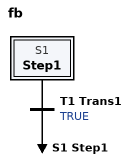
   // sequencer 1
   INITIAL_STEP Step1:   // S1, max time T#10S, warning time T#7S
   END_STEP
   TRANSITION Trans1 FROM Step1 TO Step1   // T1, jump
      := TRUE;
   END_TRANSITION
END_FUNCTION_BLOCK

ORGANIZATION_BLOCK "Main"   // OB1, LAD, ProgramCycle
TITLE = "Main Program Sweep (Cycle)"
{ S7_Optimized_Access := 'TRUE' }
VERSION : 0.1
   VAR_INPUT
      Initial_Call : Bool;   // Initial call of this OB
      Remanence : Bool;   // =True, if remanent data are available
   END_VAR
BEGIN

REGION Network 1
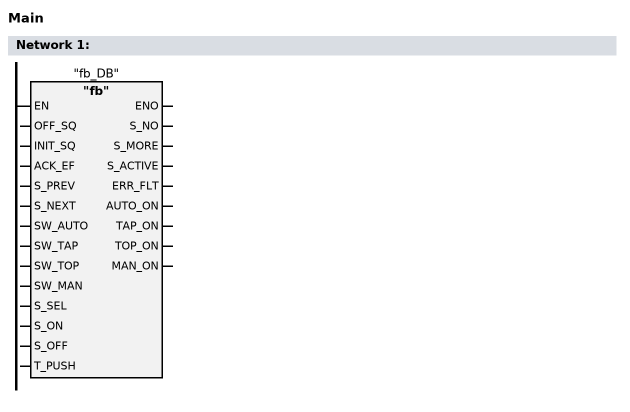
   RUNG wire#powerrail
      "fb_DB"(OFF_SQ :=, INIT_SQ :=, ACK_EF :=, S_PREV :=, S_NEXT :=, SW_AUTO :=, SW_TAP :=, SW_TOP :=, SW_MAN :=, S_SEL :=, S_ON :=, S_OFF :=, T_PUSH :=, S_NO =>, S_MORE =>, S_ACTIVE =>, ERR_FLT =>, AUTO_ON =>, TAP_ON =>, TOP_ON =>, MAN_ON =>)
   END_RUNG
   // the same network as SCL:
   "fb_DB"();   // "fb"
END_REGION
END_ORGANIZATION_BLOCK

(* ===== HMI "HMI_RT_2" =====
system functions are stored by id; their names below are inferred from use
connection "Connection_1": ETHERNET, SIMATIC S7 300/400 MPI
connection "HMI_Connection_1": ETHERNET, SIMATIC S7 300/400 MPI

HMI tags "Default tag table"
   "Tag_ScreenNumber" : UInt, internal
   "Greutate" : Int AT %DB7.DBW2, 1 s
   "LOAD" : Bool = PLC Banda_1_DB.Btn_LOAD AT %DB8.DBX0.4, 1 s
   "Manuala" : UInt, internal
   "Automata" : UInt, internal
   "StatieDistributie" : UInt, internal
   "StatieHidraulica" : UInt, internal
   "StatieIncarcare" : UInt, internal
   "Poz_Piston_1" : Int = PLC DB_general.Poz_Piston_1 AT %DB2.DBW2, 500 ms
   "Emg_Stop" : Bool = PLC Emg_Stop AT %I0.2, 1 s
   "Poz_Cutie" : Int = PLC Poz_Cutie AT %MW0, 500 ms
   "DB_general_Stare_Poz_Incarcare" : Bool = PLC DB_general.Stare_Poz_Incarcare AT %DB2.DBX0.0, 1 s
   "ON/OFF" : Bool = PLC "ON/OFF" AT %M2.1, 1 s
   "Viz_Cutie_Cursa_Scurta" : Bool = PLC Viz_Cutie_Cursa_Scurta AT %M2.2, 500 ms
   "Final_Cursa_P1" : Bool = PLC Final_Cursa_Piston_1 AT %M2.5, 1 s
   "Locuri_A" : Int = PLC DB_HMI.Locuri_A AT %DB19.DBW0, 1 s
   "Locuri_B" : Int = PLC DB_HMI.Locuri_B AT %DB19.DBW2, 1 s
   "Locuri_C" : Int = PLC DB_HMI.Locuri_C AT %DB19.DBW4, 1 s
   "Loc_Ocupat_A" : Int AT %DB1.DBW0, 1 s
   "DB_general_Poz_Piston_1" : Int = PLC DB_general.Poz_Piston_1 AT %DB2.DBW2, 1 s
   "DB_HMI_A_Pressed" : Bool = PLC DB_HMI.A_Pressed AT %DB19.DBX6.0, 1 s
   "DB_HMI_B_Pressed" : Bool = PLC DB_HMI.B_Pressed AT %DB19.DBX6.1, 1 s
   "DB_HMI_C_Pressed" : Bool = PLC DB_HMI.C_Pressed AT %DB19.DBX6.2, 1 s
   "DB_HMI_Cutie_Manuala" : Bool = PLC DB_HMI.Cutie_Manuala AT %DB19.DBX6.4, 1 s
   "DB_HMI_Cutie_Automata" : Bool = PLC DB_HMI.Cutie_Automata AT %DB19.DBX6.3, 1 s
   "DB_HMI_Viz_Cutie_Scurta" : Bool = PLC DB_HMI.Viz_Cutie_Scurta AT %DB19.DBX6.5, 1 s
   "DB_general_Senzor_1_Incarcare" : Bool = PLC DB_general.Senzor_1_Incarcare AT %DB2.DBX0.2, 1 s
   "DB_general_Senzor_2_Incarcare" : Bool = PLC DB_general.Senzor_2_Incarcare AT %DB2.DBX0.3, 1 s
   "DB_HMI_Tip_Cutie" : Int = PLC DB_HMI.Tip_Cutie_Lung AT %DB19.DBW8, 1 s
   "DB_HMI_LOAD" : Int = PLC DB_HMI.LOAD AT %DB19.DBW12, 1 s
   "DB_HMI_Transport" : Bool = PLC DB_HMI.Transport AT %DB19.DBX14.0, 1 s
   "DB_HMI_Viz_Cutie_Lunga" : Bool = PLC DB_HMI.Viz_Cutie_Lunga AT %DB19.DBX6.6, 1 s
   "DB_HMI_Tip_Cutie_Scurt" : Int = PLC DB_HMI.Tip_Cutie_Scurt AT %DB19.DBW10, 1 s
   "DB_general_Senzor_1_Descarcare" : Bool = PLC DB_general.Senzor_1_Descarcare AT %DB2.DBX0.4, 1 s
   "Stop" : Bool = PLC Stop AT %I0.1, 1 s
   "Start" : Bool = PLC Start AT %I0.0, 1 s
   "Man/Auto" : Bool = PLC "Man/Auto" AT %I0.3, 1 s
   "DB_general_Valoare" : Int = PLC DB_general.Valoare AT %DB2.DBW14, 1 s
   "DB_general_Piston_Cursa_Completa" : Int = PLC DB_general.Piston_1_Cursa_Completa AT %DB2.DBW16, 500 ms
   "DB_HMI_Viz_Cutie_Banda_1" : Bool = PLC DB_HMI.Viz_Cutie_Banda_1 AT %DB19.DBX14.2, 500 ms
   "DB_HMI_Ack_Load" : Bool = PLC DB_HMI.Ack_Load AT %DB19.DBX14.3, 1 s
   "DB_HMI_Piston_1_Status" : Int = PLC DB_HMI.Piston_1_Status AT %DB19.DBW16, 1 s
   "DB_HMI_Piston_2_Status" : Int = PLC DB_HMI.Piston_2_Status AT %DB19.DBW18, 1 s
   "DB_general_Piston_2_Cursa_Completa" : Int = PLC DB_general.Piston_2_Cursa_Completa AT %DB2.DBW18, 500 ms
   "DB_HMI_Load_RDY" : Bool = PLC DB_HMI.Load_RDY AT %DB19.DBX20.0, 1 s
   "DB_general_Poz_Cutie_Bile" : Int = PLC DB_general.Poz_Cutie_Bile AT %DB2.DBW8, 500 ms
   "DB_HMI_Viz_Cutie_A" : Bool = PLC DB_HMI.Viz_Cutie_A AT %DB19.DBX20.1, 1 s
   "DB_HMI_Viz_Cutie_B" : Bool = PLC DB_HMI.Viz_Cutie_B AT %DB19.DBX20.2, 1 s
   "DB_HMI_Viz_Cutie_C" : Bool = PLC DB_HMI.Viz_Cutie_C AT %DB19.DBX20.3, 1 s
   "DB_HMI_LOAD_A" : Bool = PLC DB_HMI.LOAD_A AT %DB19.DBX28.0, 1 s
   "DB_general_Piston_Incarcare_A" : Int = PLC DB_general.Piston_Incarcare_A AT %DB2.DBW30, 500 ms
   "DB_HMI_LOAD_B" : Bool = PLC DB_HMI.LOAD_B AT %DB19.DBX28.1, 1 s
   "DB_HMI_LOAD_C" : Bool = PLC DB_HMI.LOAD_C AT %DB19.DBX28.2, 1 s
   "DB_general_Piston_Incarcare_B" : Int = PLC DB_general.Piston_Incarcare_B AT %DB2.DBW32, 1 s
   "DB_general_Piston_Incarcare_C" : Int = PLC DB_general.Piston_Incarcare_C AT %DB2.DBW34, 1 s
   "DB_HMI_Status_Piston_A" : Int = PLC DB_HMI.Status_Piston_A AT %DB19.DBW22, 1 s
   "DB_HMI_Status_Piston_B" : Int = PLC DB_HMI.Status_Piston_B AT %DB19.DBW24, 1 s
   "DB_HMI_Status_Piston_C" : Int = PLC DB_HMI.Status_Piston_C AT %DB19.DBW26, 1 s
   "DB_HMI_Status_Banda_Bile" : Int = PLC DB_HMI.Status_Banda_Bile AT %DB19.DBW30, 1 s
   "DB_HMI_Sageata_Deplasare_Banda_Bile" : Bool = PLC DB_HMI.Sageata_Deplasare_Banda_Bile AT %DB19.DBX32.0, 1 s
   "DB_HMI_Temp_Ulei" : Int = PLC DB_HMI.Temp_Ulei AT %DB19.DBW34, 500 ms
   "DB_HMI_Volum_Ulei" : Int = PLC DB_HMI.Volum_Ulei AT %DB19.DBW40, 1 s
   "DB_HMI_Add_Ulei" : Bool = PLC DB_HMI.Add_Ulei AT %DB19.DBX42.0, 1 s
   "DB_HMI_Sub_Ulei" : Bool = PLC DB_HMI.Sub_Ulei AT %DB19.DBX42.1, 1 s
   "DB_HMI_Start_System" : Bool = PLC DB_HMI.Start_System AT %DB19.DBX42.2, 1 s
   "DB_HMI_Racire_Ulei" : Bool = PLC DB_HMI.Racire_Ulei AT %DB19.DBX42.3, 1 s
   "DB_HMI_Set_T0" : Bool = PLC DB_HMI.Set_T0 AT %DB19.DBX42.6, 1 s
   "DB_HMI_Set_T50" : Bool = PLC DB_HMI.Set_T50 AT %DB19.DBX42.7, 1 s
   "DB_HMI_START_SIM" : Bool = PLC DB_HMI.START_SIM AT %DB19.DBX43.0, 1 s
   "DB_SIM_BTN_RESET" : Bool = PLC DB_SIM.BTN_RESET AT %DB40.DBX0.4, 1 s
   "DB_HMI_TEST_LOAD" : Bool = PLC DB_HMI.BTN_LOAD AT %DB19.DBX43.1, 1 s
   "DB_Alarme_Emg_Stop" : Int = PLC DB_Alarme.Emg_Stop AT %DB46.DBW0, 1 s

discrete alarms
   1: 'Emergency Stop', class Errors, trigger "DB_Alarme_Emg_Stop" bit 0

analog alarms
   1: 'Limita greutate depasita / Gewichtslimit überschritten', class Warnings, trigger "Greutate"
   2: 'No more free spaces in A slot / Keine freien Plätze mehr im A-Steckplatz', class Acknowledgement, trigger "Locuri_A"
   3: 'No more free spaces in B slot / Keine freien Plätze mehr im B-Steckplatz', class Acknowledgement, trigger "Locuri_B"
   4: 'No more free spaces in C slot / Keine freien Plätze mehr im C-Steckplatz', class Acknowledgement, trigger "Locuri_C"
   5: 'Hydraulic oil overheated / Hydrauliköl überhitzt', class Errors, trigger "DB_HMI_Temp_Ulei"
   6: 'Hydraulic oil too cold / Hydrauliköl zu kalt', class Errors, trigger "DB_HMI_Temp_Ulei"
   7: 'Hydraulic oil volume too high / Hydraulikölmenge zu hoch', class Errors, trigger "DB_HMI_Volum_Ulei"
   8: 'Hydraulic oil volume too low / Hydraulikölmenge zu gering', class Errors, trigger "DB_HMI_Volum_Ulei"

Template "Template_1" 320x240
   Button "Exit" at 266,202 size 52x37; TextOff 'Exit / Ausfahrt'; PictureOff "ExitRuntime_KTP600_Basic_color_PN"; PictureOn "ExitRuntime_KTP600_Basic_color_PN"
      on Release: StopRuntime(0)
   Button "Template_Button" at 213,202 size 52x37; TextOff 'Text'
   Button "Template_Button_1" at 160,202 size 52x37; TextOff 'Text'
   Button "Template_Button_2" at 107,202 size 52x37; TextOff 'Text'
   Button "Template_Button_3" at 54,202 size 52x37; TextOff 'Text'
   Button "Start screen" at 1,202 size 52x37; TextOff 'Start screen / Startbildschirm'; PictureOff "NavigateHome_KTP600_Basic_color_PN"; PictureOn "NavigateHome_KTP600_Basic_color_PN"
      on Release: ActivateScreen("Home", 0)
   SymbolicIOField "Symbolic_IO_Field_Screen" at 69,7 size 164x24; TextOff '0'; TextOn '1'; TextList "TextList_ScreenNames"
      ProcessValue <- "Tag_ScreenNumber"
      on Change: ActivateScreenByNumber("Tag_ScreenNumber", 0)
   DateTimeField "HmiScreenItemData" at 235,19 size 85x19
   DateTimeField "HmiScreenItemData_1" at 235,0 size 85x19
   GraphicView "Logo" at 0,0 size 67x38; Picture "Logo of HMI_1"

screen "Home" 320x240, template "Template_2"
   on GenerateScreen: SetTag("Tag_ScreenNumber", 1)
   GraphicView "Graphic view_10" at 119,49 size 40x42; Picture "Graphic_42"
   Rectangle "Rectangle_45" at 129,65 size 24x20
      Visibility <- "DB_HMI_B_Pressed"
      VerticalMovement <- "DB_general_Poz_Cutie_Bile"
   Rectangle "Rectangle_47" at 128,65 size 25x20
      Visibility <- "DB_HMI_A_Pressed"
      VerticalMovement <- "DB_general_Poz_Cutie_Bile"
   Rectangle "Rectangle_49" at 128,65 size 25x20
      Visibility <- "DB_HMI_C_Pressed"
      VerticalMovement <- "DB_general_Poz_Cutie_Bile"
   GraphicView "Graphic view_8" at 130,66 size 21x18; Picture "Box"
      Visibility <- "DB_HMI_Viz_Cutie_A"
      VerticalMovement <- "DB_general_Poz_Cutie_Bile"
   GraphicView "Graphic view_9" at 130,66 size 21x18; Picture "Box"
      Visibility <- "DB_HMI_Viz_Cutie_B"
      VerticalMovement <- "DB_general_Poz_Cutie_Bile"
   GraphicView "Graphic view_11" at 130,66 size 21x18; Picture "Box"
      Visibility <- "DB_HMI_Viz_Cutie_C"
      VerticalMovement <- "DB_general_Poz_Cutie_Bile"
   GraphicView "Graphic view_5" at 119,20 size 40x42; Picture "Graphic_42"
   Rectangle "Rectangle_17" at 137,13 size 9x14
      VerticalMovement <- "DB_general_Piston_2_Cursa_Completa"
   Rectangle "Rectangle_18" at 135,13 size 12x14
      VerticalMovement <- "DB_general_Piston_2_Cursa_Completa"
   Rectangle "Rectangle_19" at 134,13 size 15x14
      VerticalMovement <- "DB_general_Piston_2_Cursa_Completa"
   Rectangle "Rectangle_1" at 107,165 size 14x6
      HorizontalMovement <- "DB_general_Piston_Incarcare_C"
   Rectangle "Rectangle_25" at 107,164 size 14x8
      HorizontalMovement <- "DB_general_Piston_Incarcare_C"
   Rectangle "Rectangle_26" at 108,163 size 14x10
      HorizontalMovement <- "DB_general_Piston_Incarcare_C"
   Rectangle "Rectangle_27" at 107,161 size 14x14
      HorizontalMovement <- "DB_general_Piston_Incarcare_C"
   Rectangle "Rectangle_28" at 107,132 size 14x6
      HorizontalMovement <- "DB_general_Piston_Incarcare_B"
   Rectangle "Rectangle_29" at 107,131 size 14x8
      HorizontalMovement <- "DB_general_Piston_Incarcare_B"
   Rectangle "Rectangle_30" at 108,130 size 14x10
      HorizontalMovement <- "DB_general_Piston_Incarcare_B"
   Rectangle "Rectangle_31" at 107,128 size 14x14
      HorizontalMovement <- "DB_general_Piston_Incarcare_B"
   Rectangle "Rectangle_32" at 107,99 size 14x6
      HorizontalMovement <- "DB_general_Piston_Incarcare_A"
   Rectangle "Rectangle_33" at 107,98 size 14x8
      HorizontalMovement <- "DB_general_Piston_Incarcare_A"
   Rectangle "Rectangle_34" at 108,97 size 14x10
      HorizontalMovement <- "DB_general_Piston_Incarcare_A"
   Rectangle "Rectangle_35" at 107,95 size 14x14
      HorizontalMovement <- "DB_general_Piston_Incarcare_A"
   GraphicView "Graphic view_3" at 157,88 size 79x26; Picture "Graphic_30"
   GraphicView "Graphic view_4" at 157,122 size 79x26; Picture "Graphic_30"
   GraphicView "Graphic view_6" at 158,153 size 79x26; Picture "Graphic_30"
   GraphicView "Graphic view_7" at 158,180 size 21x9; Picture "Graphic_32"
   Rectangle "Rectangle_50" at 196,92 size 14x11
      Appearance <- "Locuri_A"
   Rectangle "Rectangle_51" at 179,92 size 14x11
      Appearance <- "Locuri_A"
   Rectangle "Rectangle_52" at 163,92 size 14x11
      Appearance <- "Locuri_A"
   Rectangle "Rectangle_53" at 196,124 size 14x11
      Appearance <- "Locuri_B"
   Rectangle "Rectangle_54" at 179,124 size 14x11
      Appearance <- "Locuri_B"
   Rectangle "Rectangle_55" at 163,124 size 14x11
      Appearance <- "Locuri_B"
   Rectangle "Rectangle_56" at 196,157 size 14x11
      Appearance <- "Locuri_C"
   Rectangle "Rectangle_57" at 179,157 size 14x11
      Appearance <- "Locuri_C"
   Rectangle "Rectangle_58" at 163,157 size 14x11
      Appearance <- "Locuri_C"
   Rectangle "Rectangle_59" at 120,91 size 5x23
      HorizontalMovement <- "DB_general_Piston_Incarcare_A"
   Rectangle "Rectangle_60" at 120,123 size 5x23
      HorizontalMovement <- "DB_general_Piston_Incarcare_B"
   Rectangle "Rectangle_61" at 120,155 size 5x23
      HorizontalMovement <- "DB_general_Piston_Incarcare_C"
   GraphicView "Graphic view_1" at 13,54 size 40x44; Picture "Graphic_42"
   Rectangle "Rectangle_8" at 32,84 size 11x13
      VerticalMovement <- "DB_general_Piston_Cursa_Completa"
   Rectangle "Rectangle_7" at 31,81 size 12x14
      VerticalMovement <- "DB_general_Piston_Cursa_Completa"
   Rectangle "Rectangle_6" at 30,81 size 15x14
      VerticalMovement <- "DB_general_Piston_Cursa_Completa"
   Rectangle "Rectangle_10" at 24,81 size 27x4
      VerticalMovement <- "DB_general_Piston_Cursa_Completa"
   GraphicView "Graphic view_2" at 26,30 size 21x23; Picture "Box"
      Visibility <- "DB_HMI_Viz_Cutie_Banda_1"
      HorizontalMovement <- "Poz_Cutie"
   TextField "Text field_8" at 60,69 size 15x13; Text 'S1'
   TextField "Text field_9" at 60,78 size 15x13; Text 'S2'
   Rectangle "Rectangle_9" at 52,72 size 7x6
      Appearance <- "DB_general_Senzor_1_Incarcare"
   Rectangle "Rectangle_14" at 52,81 size 7x6
      Appearance <- "DB_general_Senzor_2_Incarcare"
   Rectangle "Rectangle_15" at 154,30 size 7x6
      Appearance <- "DB_general_Senzor_1_Descarcare"
   Rectangle "Rectangle_16" at 154,40 size 7x6
      Appearance <- "DB_general_Senzor_1_Descarcare"
   TextField "Text field_13" at 163,37 size 15x13; Text 'S4'
   Rectangle "Rectangle_21" at 128,26 size 25x4
      VerticalMovement <- "DB_general_Piston_2_Cursa_Completa"
   TextField "Text field_1" at 163,27 size 15x13; Text 'S3'

screen "StatieIncarcare" 320x240, template "Template_2"
   GraphicView "Graphic view_10" at 26,0 size 48x44; Picture "background.xwr"
   Rectangle "Rectangle_15" at 32,6 size 39x32
      VerticalMovement <- "DB_general_Poz_Cutie_Bile"
      Visibility <- "DB_HMI_B_Pressed"
   Rectangle "Rectangle_24" at 32,6 size 40x32
      Visibility <- "DB_HMI_A_Pressed"
      VerticalMovement <- "DB_general_Poz_Cutie_Bile"
   Rectangle "Rectangle_16" at 32,5 size 40x33
      VerticalMovement <- "DB_general_Poz_Cutie_Bile"
      Visibility <- "DB_HMI_C_Pressed"
   Switch "Switch_1" at 83,7 size 71x24; CaptionText 'Switch'; TextOff 'Transport'; TextOn 'Transporting / Transport'
      ProcessValue <- "DB_HMI_Transport"
      Appearance <- "DB_HMI_Transport"
   Switch "Switch_2" at 252,47 size 63x28; CaptionText 'Switch'; TextOff 'LOAD A BELASTUNG A'; TextOn 'LOADIGN A LADEN A'
      ProcessValue <- "DB_HMI_LOAD_A"
      Appearance <- "DB_HMI_A_Pressed"
   Switch "Switch_3" at 253,91 size 63x28; TextOn 'LOADIGN B LADEN B'; CaptionText 'Switch'; TextOff 'LOAD B BELASTUNG B'
      ProcessValue <- "DB_HMI_LOAD_B"
      Appearance <- "DB_HMI_B_Pressed"
   Switch "Switch_4" at 254,135 size 63x28; TextOn 'LOADIGN C LADEN C'; CaptionText 'Switch'; TextOff 'LOAD C BELASTUNG C'
      ProcessValue <- "DB_HMI_LOAD_C"
      Appearance <- "DB_HMI_C_Pressed"
   GraphicView "Graphic view_8" at 136,188 size 21x18; Picture "Graphic_43"
      Visibility <- "DB_HMI_Sageata_Deplasare_Banda_Bile"
   GraphicView "Graphic view_9" at 112,188 size 21x18; Picture "Graphic_44"
      Visibility <- "DB_HMI_Sageata_Deplasare_Banda_Bile"
   GraphicIOField "PlotLight_Round_G" at 253,183 size 23x22; PictureOff "PilotLight_Round_G_Off_256c"; PictureOn "PilotLight_Round_G_On_256c"
      ProcessValue <- "ON/OFF"
   GraphicIOField "PlotLight_Round_R" at 230,182 size 23x22; PictureOff "PilotLight_Round_R_On_256c"; PictureOn "PilotLight_Round_R_Off_256c"
      ProcessValue <- "ON/OFF"
   Switch "Rotary_N" at 278,182 size 34x25; CaptionText 'Switch'; TextOff '0'; TextOn '1'; PictureOff "Rotary_N_On_256c"; PictureOn "Rotary_N_Off_256c"
      ProcessValue <- "Man/Auto"
   TextField "Text field_4" at 230,172 size 20x10; Text 'STOP'
   TextField "Text field_5" at 252,172 size 24x10; Text 'START'
   TextField "Text field_6" at 275,173 size 18x10; Text 'MAN'
   TextField "Text field_7" at 295,173 size 21x10; Text 'AUTO'
   Rectangle "Rectangle_6" at 0,164 size 21x10
      HorizontalMovement <- "DB_general_Piston_Incarcare_C"
   Rectangle "Rectangle_7" at 0,163 size 21x12
      HorizontalMovement <- "DB_general_Piston_Incarcare_C"
   Rectangle "Rectangle_8" at 1,161 size 21x16
      HorizontalMovement <- "DB_general_Piston_Incarcare_C"
   Rectangle "Rectangle_10" at 0,158 size 21x22
      HorizontalMovement <- "DB_general_Piston_Incarcare_C"
   Rectangle "Rectangle_3" at 0,112 size 21x10
      HorizontalMovement <- "DB_general_Piston_Incarcare_B"
   Rectangle "Rectangle_4" at 0,111 size 21x12
      HorizontalMovement <- "DB_general_Piston_Incarcare_B"
   Rectangle "Rectangle_5" at 1,109 size 21x16
      HorizontalMovement <- "DB_general_Piston_Incarcare_B"
   Rectangle "Rectangle_17" at 0,106 size 21x22
      HorizontalMovement <- "DB_general_Piston_Incarcare_B"
   Rectangle "Rectangle_30" at 0,60 size 21x10
      HorizontalMovement <- "DB_general_Piston_Incarcare_A"
   Rectangle "Rectangle_29" at 0,59 size 21x12
      HorizontalMovement <- "DB_general_Piston_Incarcare_A"
   Rectangle "Rectangle_28" at 1,57 size 21x16
      HorizontalMovement <- "DB_general_Piston_Incarcare_A"
   Rectangle "Rectangle_25" at 0,54 size 21x22
      HorizontalMovement <- "DB_general_Piston_Incarcare_A"
   GraphicView "Graphic view_3" at 75,43 size 119x41; Picture "Graphic_30"
   GraphicView "Graphic view_2" at 75,96 size 119x41; Picture "Graphic_30"
   GraphicView "Graphic view_4" at 76,145 size 119x41; Picture "Graphic_30"
   Button "Button_2" at 194,179 size 37x25; TextOff 'EMG STOP EMG STOP'
      on Press: SetTag("Emg_Stop", 0)
      Appearance <- "Emg_Stop"
      Visibility <- "Emg_Stop"
   Rectangle "Rectangle_48" at 5,85 size 20x13
      Appearance <- "DB_HMI_Status_Piston_A"
   TextField "Text field_8" at 5,83 size 21x13; Text 'P-A'
   GraphicView "Graphic view_5" at 77,190 size 31x15; Picture "Graphic_32"
   Rectangle "Rectangle_9" at 133,50 size 21x17
      Appearance <- "Locuri_A"
   Rectangle "Rectangle_13" at 108,50 size 21x17
      Appearance <- "Locuri_A"
   Rectangle "Rectangle_14" at 83,50 size 21x17
      Appearance <- "Locuri_A"
   Rectangle "Rectangle_18" at 133,101 size 21x17
      Appearance <- "Locuri_B"
   Rectangle "Rectangle_19" at 108,101 size 21x17
      Appearance <- "Locuri_B"
   Rectangle "Rectangle_20" at 83,101 size 21x17
      Appearance <- "Locuri_B"
   Rectangle "Rectangle_21" at 133,153 size 21x17
      Appearance <- "Locuri_C"
   Rectangle "Rectangle_22" at 108,153 size 21x17
      Appearance <- "Locuri_C"
   Rectangle "Rectangle_23" at 83,153 size 21x17
      Appearance <- "Locuri_C"
   GraphicView "Graphic view_1" at 35,7 size 32x29; Picture "Box"
      VerticalMovement <- "DB_general_Poz_Cutie_Bile"
      Visibility <- "DB_HMI_Viz_Cutie_A"
   Rectangle "Rectangle_27" at 19,47 size 7x37
      HorizontalMovement <- "DB_general_Piston_Incarcare_A"
   Rectangle "Rectangle_32" at 19,99 size 7x37
      HorizontalMovement <- "DB_general_Piston_Incarcare_B"
   Rectangle "Rectangle_12" at 19,151 size 7x37
      HorizontalMovement <- "DB_general_Piston_Incarcare_C"
   GraphicView "Graphic view_7" at 36,6 size 32x29; Picture "Box"
      Visibility <- "DB_HMI_Viz_Cutie_B"
      VerticalMovement <- "DB_general_Poz_Cutie_Bile"
   GraphicView "Graphic view_6" at 36,7 size 32x29; Picture "Box"
      Visibility <- "DB_HMI_Viz_Cutie_C"
      VerticalMovement <- "DB_general_Poz_Cutie_Bile"
   Rectangle "Rectangle_33" at 85,194 size 14x7
      Appearance <- "DB_HMI_Status_Banda_Bile"
   Rectangle "Rectangle_49" at 6,137 size 20x13
      Appearance <- "DB_HMI_Status_Piston_B"
   Rectangle "Rectangle_50" at 6,190 size 20x13
      Appearance <- "DB_HMI_Status_Piston_C"
   TextField "Text field_11" at 6,135 size 20x13; Text 'P-B'
   TextField "Text field_9" at 6,188 size 20x13; Text 'P-C'

screen "Animatie_B1" 320x240, template "Template_2"
   GraphicIOField "PlotLight_Round_G" at 242,177 size 27x25; PictureOn "PilotLight_Round_G_On_256c"; PictureOff "PilotLight_Round_G_Off_256c"
      ProcessValue <- "ON/OFF"
   GraphicIOField "PlotLight_Round_R" at 215,176 size 27x25; PictureOn "PilotLight_Round_R_Off_256c"; PictureOff "PilotLight_Round_R_On_256c"
      ProcessValue <- "ON/OFF"
   Switch "Rotary_N" at 272,176 size 41x29; CaptionText 'Switch'; TextOff '0'; TextOn '1'; PictureOn "Rotary_N_Off_256c"; PictureOff "Rotary_N_On_256c"
      ProcessValue <- "Man/Auto"
   TextField "Text field_4" at 220,167 size 20x10; Text 'STOP'
   TextField "Text field_5" at 244,167 size 24x10; Text 'START'
   TextField "Text field_6" at 268,165 size 18x10; Text 'MAN'
   TextField "Text field_7" at 292,165 size 21x10; Text 'AUTO'
   Button "Button_2" at 176,172 size 39x29; TextOff 'EMG STOP EMG STOP'
      on Press: SetTag("Emg_Stop", 0)
      Appearance <- "Emg_Stop"
      Visibility <- "Emg_Stop"
   Switch "Switch_6" at 0,181 size 45x28; TextOn 'Placed Box Kolben Status'; CaptionText 'Switch'; TextOff 'Place Box Kolben Status'
      on SwitchOff: SetTag("DB_general_Senzor_1_Incarcare", 0); SetTag("DB_general_Senzor_2_Incarcare", 0)
      on SwitchOn: SetTag("DB_general_Senzor_1_Incarcare", 1); SetTag("DB_general_Senzor_2_Incarcare", 1)
      Appearance <- "DB_HMI_Viz_Cutie_Scurta"
      ProcessValue <- "DB_HMI_Viz_Cutie_Scurta"
   Switch "Switch_1" at 47,181 size 45x28; TextOn 'ACK LOAD ACK LAST'; CaptionText 'Switch'; TextOff 'ACK LOAD ACK LAST'
      Appearance <- "DB_general_Stare_Poz_Incarcare"
      ProcessValue <- "DB_HMI_Ack_Load"
      on SwitchOn: SetTag("DB_HMI_Load_RDY", 1)
   Group "Group" at 172,163 size 143x45; PictureOff "PilotLight_Round_G_Off_256c"; PictureOn "PilotLight_Round_G_On_256c"
   Switch "Switch_8" at 251,126 size 64x32; TextOn 'Started Sim / Sim gestartet'; CaptionText 'Switch'; TextOff 'Start Sim / Starten Sie Sim'
      ProcessValue <- "DB_HMI_START_SIM"
      Appearance <- "DB_HMI_START_SIM"
   IOField "I/O field_1" at 281,44 size 33x15; FormatPattern 99
      ProcessValue <- "Poz_Cutie"
   Switch "Switch_2" at 94,181 size 45x28; CaptionText 'Switch'; TextOff 'LOAD / BELASTUNG'; TextOn 'LOAD / BELASTUNG'
      ProcessValue <- "DB_HMI_TEST_LOAD"
      Appearance <- "DB_HMI_TEST_LOAD"
   Button "Button_1" at 256,91 size 55x32; TextOff 'RESET / ZURÜCKSETZEN'
      on Press: SetTag("DB_HMI_Viz_Cutie_Scurta", 0); SetTag("LOAD", 0); SetTag("DB_HMI_Ack_Load", 0); SetTag("DB_SIM_BTN_RESET", 1); SetTag("DB_general_Senzor_1_Incarcare", 0); SetTag("DB_general_Senzor_2_Incarcare", 0); SetTag("LOAD", 0); SetTag("DB_HMI_TEST_LOAD", 0)
      on Release: SetTag("DB_SIM_BTN_RESET", 0)
   IOField "I/O field_2" at 124,133 size 19x15; FormatPattern 9
      ProcessValue <- "Locuri_A"
   IOField "I/O field_3" at 166,133 size 19x15; FormatPattern 9
      ProcessValue <- "Locuri_B"
   IOField "I/O field_4" at 209,133 size 19x15; FormatPattern 9
      ProcessValue <- "Locuri_C"
   Switch "Switch_3" at 120,105 size 27x23; TextOn 'A'; CaptionText 'Switch'; TextOff 'A'
      on SwitchOff: SetTag("DB_HMI_Viz_Cutie_A", 0)
      on SwitchOn: SetTag("DB_HMI_B_Pressed", 0); SetTag("DB_HMI_C_Pressed", 0); SetTag("DB_HMI_Viz_Cutie_A", 1); SetTag("DB_HMI_Viz_Cutie_B", 0); SetTag("DB_HMI_Viz_Cutie_C", 0)
      Appearance <- "DB_HMI_A_Pressed"
      ProcessValue <- "DB_HMI_A_Pressed"
   Switch "Switch_4" at 162,104 size 27x23; TextOn 'B'; CaptionText 'Switch'; TextOff 'B'
      on SwitchOn: SetTag("DB_HMI_A_Pressed", 0); SetTag("DB_HMI_C_Pressed", 0); SetTag("DB_HMI_Viz_Cutie_B", 1); SetTag("DB_HMI_Viz_Cutie_A", 0); SetTag("DB_HMI_Viz_Cutie_C", 0)
      Appearance <- "DB_HMI_B_Pressed"
      ProcessValue <- "DB_HMI_B_Pressed"
   Switch "Switch_5" at 204,104 size 27x23; TextOn 'C'; CaptionText 'Switch'; TextOff 'C'
      on SwitchOn: SetTag("DB_HMI_A_Pressed", 0); SetTag("DB_HMI_B_Pressed", 0); SetTag("DB_HMI_Viz_Cutie_C", 1); SetTag("DB_HMI_Viz_Cutie_B", 0); SetTag("DB_HMI_Viz_Cutie_A", 0)
      Appearance <- "DB_HMI_C_Pressed"
      ProcessValue <- "DB_HMI_C_Pressed"
   IOField "I/O field_5" at 0,145 size 24x15; FormatPattern 99
      ProcessValue <- "DB_general_Piston_Cursa_Completa"
   IOField "I/O field_6" at 191,0 size 33x15; FormatPattern 99
      ProcessValue <- "DB_general_Piston_2_Cursa_Completa"
   Rectangle "Rectangle_25" at 233,4 size 15x13
      Appearance <- "DB_HMI_Piston_2_Status"
   TextField "Text field_3" at 233,3 size 16x13; Text 'P2'
   GraphicView "Graphic view_5" at 191,30 size 65x62; Picture "Graphic_42"
   Rectangle "Rectangle_17" at 220,19 size 17x20
      VerticalMovement <- "DB_general_Piston_2_Cursa_Completa"
   Rectangle "Rectangle_18" at 218,19 size 20x20
      VerticalMovement <- "DB_general_Piston_2_Cursa_Completa"
   Rectangle "Rectangle_19" at 216,19 size 24x21
      VerticalMovement <- "DB_general_Piston_2_Cursa_Completa"
   Rectangle "Rectangle_24" at 34,145 size 15x13
      Appearance <- "DB_HMI_Piston_1_Status"
   TextField "Text field_2" at 34,144 size 16x13; Text 'P1'
   GraphicView "Graphic view_1" at 20,80 size 65x64; Picture "Graphic_42"
   Rectangle "Rectangle_8" at 51,124 size 17x20
      VerticalMovement <- "DB_general_Piston_Cursa_Completa"
   Rectangle "Rectangle_7" at 50,120 size 20x20
      VerticalMovement <- "DB_general_Piston_Cursa_Completa"
   Rectangle "Rectangle_6" at 48,120 size 24x21
      VerticalMovement <- "DB_general_Piston_Cursa_Completa"
   Rectangle "Rectangle_10" at 38,120 size 43x6
      VerticalMovement <- "DB_general_Piston_Cursa_Completa"
   GraphicView "Graphic view_2" at 42,45 size 34x34; Picture "Box"
      Visibility <- "DB_HMI_Viz_Cutie_Banda_1"
      HorizontalMovement <- "Poz_Cutie"
   TextField "Text field_8" at 97,102 size 15x13; Text 'S1'
   TextField "Text field_9" at 97,115 size 15x13; Text 'S2'
   Rectangle "Rectangle_9" at 83,106 size 11x9
      Appearance <- "DB_general_Senzor_1_Incarcare"
   Rectangle "Rectangle_14" at 83,120 size 11x9
      Appearance <- "DB_general_Senzor_2_Incarcare"
   Rectangle "Rectangle_15" at 249,45 size 11x9
      Appearance <- "DB_general_Senzor_1_Descarcare"
   Rectangle "Rectangle_16" at 249,59 size 11x9
      Appearance <- "DB_general_Senzor_1_Descarcare"
   TextField "Text field_13" at 263,54 size 15x13; Text 'S4'
   Rectangle "Rectangle_21" at 206,38 size 41x6
      VerticalMovement <- "DB_general_Piston_2_Cursa_Completa"
   TextField "Text field_1" at 262,40 size 15x13; Text 'S3'
   GraphicView "Graphic view_3" at 36,9 size 42x20; Picture "Graphic_32"
   GraphicView "Graphic view_4" at 146,9 size 42x20; Picture "Graphic_32"
   Rectangle "Rectangle_22" at 46,12 size 19x11
      Appearance <- "Poz_Cutie"
   TextField "Text field_10" at 46,9 size 18x13; Text 'M1'
   Rectangle "Rectangle_23" at 158,12 size 20x11
      Appearance <- "Poz_Cutie"
   TextField "Text field_11" at 160,9 size 18x13; Text 'M2'

screen "StatieDistribuire" 320x240, template "Template_2"
   GraphicIOField "PlotLight_Round_G" at 246,182 size 23x21; PictureOff "PilotLight_Round_G_Off_256c"; PictureOn "PilotLight_Round_G_On_256c"
      ProcessValue <- "ON/OFF"
   GraphicIOField "PlotLight_Round_R" at 221,182 size 23x21; PictureOff "PilotLight_Round_R_On_256c"; PictureOn "PilotLight_Round_R_Off_256c"
      ProcessValue <- "ON/OFF"
   Switch "Rotary_N" at 276,182 size 36x24; CaptionText 'Switch'; TextOff '0'; TextOn '1'; PictureOff "Rotary_N_On_256c"; PictureOn "Rotary_N_Off_256c"
      ProcessValue <- "Man/Auto"
   TextField "Text field_14" at 221,170 size 20x10; Text 'STOP'
   TextField "Text field_15" at 244,170 size 24x10; Text 'START'
   TextField "Text field_16" at 269,170 size 18x10; Text 'MAN'
   TextField "Text field_17" at 293,169 size 21x10; Text 'AUTO'
   Button "Button_2" at 186,184 size 30x22; TextOff 'EMG STOP EMG STOP'
      on Press: SetTag("Emg_Stop", 0)
      Appearance <- "Emg_Stop"
      Visibility <- "Emg_Stop"
   GraphicView "Graphic view_5" at 147,86 size 56x45; Picture "Graphic_42"
   Rectangle "Rectangle_17" at 174,79 size 9x15
      VerticalMovement <- "DB_general_Piston_2_Cursa_Completa"
   Rectangle "Rectangle_18" at 171,79 size 15x15
      VerticalMovement <- "DB_general_Piston_2_Cursa_Completa"
   Rectangle "Rectangle_19" at 168,79 size 21x15
      VerticalMovement <- "DB_general_Piston_2_Cursa_Completa"
   GraphicView "Graphic view_1" at 1,124 size 56x47; Picture "Graphic_42"
   Rectangle "Rectangle_8" at 28,156 size 13x15
      VerticalMovement <- "DB_general_Piston_Cursa_Completa"
   Rectangle "Rectangle_7" at 26,156 size 17x15
      VerticalMovement <- "DB_general_Piston_Cursa_Completa"
   Rectangle "Rectangle_6" at 24,156 size 21x15
      VerticalMovement <- "DB_general_Piston_Cursa_Completa"
   IOField "I/O field_1" at 10,16 size 45x25; FormatPattern 99999
      ProcessValue <- "Greutate"
   TextField "Text field_1" at 9,0 size 41x13; Text 'Weight / Gewicht'
   TextField "Text field_2" at 92,0 size 69x13; Text 'Gearbox type'
   IOField "I/O field_2" at 208,56 size 19x15; FormatPattern 9
      ProcessValue <- "Locuri_A"
   IOField "I/O field_3" at 250,56 size 19x15; FormatPattern 9
      ProcessValue <- "Locuri_B"
   IOField "I/O field_4" at 292,56 size 19x15; FormatPattern 9
      ProcessValue <- "Locuri_C"
   TextField "Text field_3" at 111,54 size 93x13; Text 'Available places / Verfügbare Plätze'
   Switch "Switch_1" at 204,28 size 27x23; CaptionText 'Switch'; TextOff 'A'; TextOn 'A'
      ProcessValue <- "DB_HMI_A_Pressed"
      Appearance <- "DB_HMI_A_Pressed"
      on SwitchOn: SetTag("DB_HMI_B_Pressed", 0); SetTag("DB_HMI_C_Pressed", 0); SetTag("DB_HMI_Viz_Cutie_A", 1); SetTag("DB_HMI_Viz_Cutie_B", 0); SetTag("DB_HMI_Viz_Cutie_C", 0)
      on SwitchOff: SetTag("DB_HMI_Viz_Cutie_A", 0)
   Switch "Switch_3" at 246,27 size 27x23; TextOn 'B'; CaptionText 'Switch'; TextOff 'B'
      ProcessValue <- "DB_HMI_B_Pressed"
      Appearance <- "DB_HMI_B_Pressed"
      on SwitchOn: SetTag("DB_HMI_A_Pressed", 0); SetTag("DB_HMI_C_Pressed", 0); SetTag("DB_HMI_Viz_Cutie_B", 1); SetTag("DB_HMI_Viz_Cutie_A", 0); SetTag("DB_HMI_Viz_Cutie_C", 0)
   Switch "Switch_4" at 288,27 size 27x23; TextOn 'C'; CaptionText 'Switch'; TextOff 'C'
      ProcessValue <- "DB_HMI_C_Pressed"
      on SwitchOn: SetTag("DB_HMI_A_Pressed", 0); SetTag("DB_HMI_B_Pressed", 0); SetTag("DB_HMI_Viz_Cutie_C", 1); SetTag("DB_HMI_Viz_Cutie_B", 0); SetTag("DB_HMI_Viz_Cutie_A", 0)
      Appearance <- "DB_HMI_C_Pressed"
   Switch "Switch_2" at 60,16 size 58x26; CaptionText 'Switch'; TextOff 'Manuala'; TextOn 'Manuala'
      ProcessValue <- "DB_HMI_Cutie_Manuala"
      Appearance <- "DB_HMI_Cutie_Manuala"
      on SwitchOn: SetTag("DB_HMI_Cutie_Automata", 0)
   Switch "Switch_5" at 134,16 size 58x26; CaptionText 'Switch'; TextOff 'Automata / Automatikgetriebe'; TextOn 'Automata / Automatikgetriebe'
      ProcessValue <- "DB_HMI_Cutie_Automata"
      Appearance <- "DB_HMI_Cutie_Automata"
      on SwitchOn: SetTag("DB_HMI_Cutie_Manuala", 0)
   Group "Group" at 182,169 size 133x40; PictureOff "PilotLight_Round_G_Off_256c"; PictureOn "PilotLight_Round_G_On_256c"
   Switch "Switch_8" at 248,135 size 61x21; CaptionText 'Switch'; TextOff 'Start Sim / Starten Sie Sim'; TextOn 'Started Sim / Sim gestartet'
      ProcessValue <- "DB_HMI_START_SIM"
      Appearance <- "DB_HMI_START_SIM"
      Visibility <- "Man/Auto"
   Switch "Switch_6" at 0,181 size 45x28; TextOn 'Placed Box Kolben Status'; CaptionText 'Switch'; TextOff 'Place Box Kolben Status'
      on SwitchOff: SetTag("DB_general_Senzor_1_Incarcare", 0); SetTag("DB_general_Senzor_2_Incarcare", 0)
      on SwitchOn: SetTag("DB_general_Senzor_1_Incarcare", 1); SetTag("DB_general_Senzor_2_Incarcare", 1)
      Appearance <- "DB_HMI_Viz_Cutie_Scurta"
      ProcessValue <- "DB_HMI_Viz_Cutie_Scurta"
   Switch "Switch_7" at 47,181 size 45x28; TextOn 'ACK LOAD ACK LAST'; CaptionText 'Switch'; TextOff 'ACK LOAD ACK LAST'
      on SwitchOn: SetTag("DB_HMI_Load_RDY", 1)
      Appearance <- "DB_general_Stare_Poz_Incarcare"
      ProcessValue <- "DB_HMI_Ack_Load"
   Switch "Switch_9" at 94,181 size 45x28; TextOn 'LOAD / BELASTUNG'; CaptionText 'Switch'; TextOff 'LOAD / BELASTUNG'
      ProcessValue <- "DB_HMI_TEST_LOAD"
      Appearance <- "DB_HMI_TEST_LOAD"
   Rectangle "Rectangle_10" at 16,153 size 37x4
      VerticalMovement <- "DB_general_Piston_Cursa_Completa"
   GraphicView "Graphic view_2" at 20,98 size 29x25; Picture "Box"
      Visibility <- "DB_HMI_Viz_Cutie_Banda_1"
      HorizontalMovement <- "Poz_Cutie"
   TextField "Text field_8" at 67,140 size 15x13; Text 'S1'
   TextField "Text field_9" at 69,149 size 15x13; Text 'S2'
   Rectangle "Rectangle_14" at 55,143 size 9x7
      Appearance <- "DB_general_Senzor_1_Incarcare"
   Rectangle "Rectangle_15" at 55,153 size 9x7
      Appearance <- "DB_general_Senzor_2_Incarcare"
   Rectangle "Rectangle_16" at 197,98 size 9x7
      Appearance <- "DB_general_Senzor_1_Descarcare"
   Rectangle "Rectangle_20" at 197,109 size 9x7
      Appearance <- "DB_general_Senzor_1_Descarcare"
   TextField "Text field_13" at 209,105 size 15x13; Text 'S4'
   Rectangle "Rectangle_22" at 160,93 size 35x4
      VerticalMovement <- "DB_general_Piston_2_Cursa_Completa"
   TextField "Text field_5" at 208,95 size 15x13; Text 'S3'
   Rectangle "Rectangle_26" at 207,75 size 15x13
      Appearance <- "DB_HMI_Piston_2_Status"
   TextField "Text field_6" at 207,74 size 16x13; Text 'P2'
   Rectangle "Rectangle_24" at 0,169 size 15x13
      Appearance <- "DB_HMI_Piston_1_Status"
   TextField "Text field_4" at 0,168 size 16x13; Text 'P1'
   GraphicView "Graphic view_3" at 6,66 size 42x20; Picture "Graphic_32"
   GraphicView "Graphic view_4" at 116,66 size 42x20; Picture "Graphic_32"
   Rectangle "Rectangle_23" at 16,69 size 19x11
      Appearance <- "Poz_Cutie"
   TextField "Text field_10" at 16,66 size 18x13; Text 'M1'
   Rectangle "Rectangle_25" at 128,69 size 20x11
      Appearance <- "Poz_Cutie"
   TextField "Text field_11" at 130,66 size 18x13; Text 'M2'
   Button "Button_1" at 248,111 size 61x21; TextOff 'RESET / ZURÜCKSETZEN'
      on Release: SetTag("DB_SIM_BTN_RESET", 0)
      on Press: SetTag("DB_HMI_Viz_Cutie_Scurta", 0); SetTag("LOAD", 0); SetTag("DB_HMI_Ack_Load", 0); SetTag("DB_SIM_BTN_RESET", 1); SetTag("DB_general_Senzor_1_Incarcare", 0); SetTag("DB_general_Senzor_2_Incarcare", 0); SetTag("LOAD", 0); SetTag("DB_HMI_TEST_LOAD", 0)
      Visibility <- "Man/Auto"
   TextField "Text field_7" at 28,100 size 15x20; Text 'M'
      Visibility <- "DB_HMI_Tip_Cutie"
      HorizontalMovement <- "Poz_Cutie"
   TextField "Text field_12" at 29,100 size 12x20; Text 'A'
      Visibility <- "DB_HMI_Tip_Cutie"
      HorizontalMovement <- "Poz_Cutie"

Template "Template_2" 320x240
   Button "Exit" at 276,209 size 38x28; TextOn 'Exit / Ausfahrt'; TextOff 'Exit / Ausfahrt'; PictureOn "ExitRuntime_KTP600_Basic_color_PN"; PictureOff "ExitRuntime_KTP600_Basic_color_PN"
      on Release: StopRuntime(0)
   Button "Template_Button_3" at 39,209 size 38x28; TextOff 'Text'
      on Press: ActivateScreen("StatieDistribuire", 4)
   Button "Start screen" at 0,209 size 38x28; TextOn 'Start screen / Startbildschirm'; TextOff 'Start screen / Startbildschirm'; PictureOn "NavigateHome_KTP600_Basic_color_PN"; PictureOff "NavigateHome_KTP600_Basic_color_PN"
      on Release: ActivateScreen("Home", 0)
   GraphicView "Logo" at 272,0 size 48x26; Picture "Logo of HMI_1"
   Button "Template_Button_1" at 78,209 size 38x28; TextOff 'Text'
      on Press: ActivateScreen("Animatie_B1", 3)
   Button "Template_Button_2" at 118,209 size 38x28; TextOff 'Text'
      on Press: ActivateScreen("Hidraulic", 0)
   Button "Template_Button_4" at 157,209 size 38x28; TextOff 'Text'
      on Press: ActivateScreen("StatieIncarcare", 0)
   Button "Template_Button_5" at 236,209 size 38x28; TextOff 'Text'
      on Press: ActivateScreen("Alarme", 0)
   GraphicView "Template_Graphic view_1" at 244,210 size 21x22; Picture "Graphic_7"
   Button "Template_Button_6" at 197,209 size 38x28; TextOff 'Text'; PictureOff "Left_Arrow"
      on Press: function_efd93a16()
   TextField "Template_Text field_1" at 41,213 size 35x13; Text 'Distrib'
   TextField "Template_Text field_2" at 82,213 size 34x13; Text 'Anima'
   TextField "Template_Text field_4" at 159,214 size 34x13; Text 'Incarc'
   TextField "Template_Text field_3" at 124,214 size 30x13; Text 'Hidra'

screen "Alarme" 320x240, template "Template_2"
   AlarmView "Alarm view_1" at 0,0 size 320x96
   SysDiagControl "System diagnostics view_1" at 1,106 size 319x96

screen "Hidraulic" 320x240, template "Template_2"
   Bar "Bar_1" at 4,16 size 54x103; Unit L; MinimumValue 0; MaximumValue 50
      ProcessValue <- "DB_HMI_Volum_Ulei"
   IOField "I/O field_1" at 27,2 size 26x19; FormatPattern 99
      ProcessValue <- "DB_HMI_Volum_Ulei"
      Appearance <- "DB_HMI_Volum_Ulei"
   Button "Button_1" at 58,40 size 23x21; TextOff '+'
      on Press: SetTag("DB_HMI_Add_Ulei", 1)
      on Release: SetTag("DB_HMI_Add_Ulei", 0)
      Appearance <- "DB_HMI_Volum_Ulei"
   Rectangle "Rectangle_1" at 57,23 size 28x15
      Appearance <- "DB_HMI_Volum_Ulei"
   Rectangle "Rectangle_2" at 56,96 size 28x15
      Appearance <- "DB_HMI_Volum_Ulei"
   TextField "Text field_1" at 58,96 size 23x13; Text 'MIN'
      Appearance <- "DB_HMI_Volum_Ulei"
   TextField "Text field_2" at 58,22 size 26x13; Text 'MAX'
      Appearance <- "DB_HMI_Volum_Ulei"
   Button "Button_2" at 58,70 size 23x21; TextOff 'Text'
      on Release: SetTag("DB_HMI_Sub_Ulei", 0)
      on Press: SetTag("DB_HMI_Sub_Ulei", 1)
      Appearance <- "DB_HMI_Volum_Ulei"
   Bar "Bar_2" at 120,17 size 54x103; Unit C; MinimumValue 0; MaximumValue 50
      ProcessValue <- "DB_HMI_Temp_Ulei"
   TextField "Text field_3" at 20,119 size 55x13; Text 'Volum Ulei / Ölvolumen'
   TextField "Text field_4" at 111,119 size 90x13; Text 'Temperatura Ulei'
   Switch "Switch_1" at 182,84 size 56x27; CaptionText 'Switch'; TextOff 'Start System Start Syst'; TextOn 'Starting System Beginnend Syst'
      ProcessValue <- "DB_HMI_Start_System"
   IOField "I/O field_3" at 145,2 size 27x20; FormatPattern 99
      ProcessValue <- "DB_HMI_Temp_Ulei"
      Appearance <- "DB_HMI_Temp_Ulei"
   GraphicView "Graphic view_2" at 182,9 size 60x53; Picture "Graphic_62"
   Rectangle "Rectangle_3" at 195,48 size 29x9
      Appearance <- "DB_HMI_Racire_Ulei"
      Visibility <- "DB_HMI_Start_System"
   TextField "Text field_7" at 6,154 size 79x13; Text 'Status Pistoane / Motorstatus'
   Rectangle "Rectangle_24" at 96,170 size 15x13
      Appearance <- "DB_HMI_Piston_1_Status"
   TextField "Text field_5" at 96,169 size 16x13; Text 'P1'
   Rectangle "Rectangle_25" at 113,170 size 15x13
      Appearance <- "DB_HMI_Piston_2_Status"
   TextField "Text field_6" at 113,170 size 16x13; Text 'P2'
   Rectangle "Rectangle_34" at 93,187 size 20x13
      Appearance <- "DB_HMI_Status_Piston_A"
   TextField "Text field_8" at 93,185 size 21x13; Text 'P-A'
   Rectangle "Rectangle_35" at 119,187 size 20x13
      Appearance <- "DB_HMI_Status_Piston_B"
   Rectangle "Rectangle_36" at 144,187 size 20x13
      Appearance <- "DB_HMI_Status_Piston_C"
   TextField "Text field_11" at 119,185 size 20x13; Text 'P-B'
   TextField "Text field_9" at 144,185 size 20x13; Text 'P-C'
   TextField "Text field_10" at 6,167 size 90x13; Text 'Statie Distribuire: / Verteilerstation:'
   TextField "Text field_12" at 4,185 size 86x13; Text 'Statie Incarcare: / Ladestation:'
   Rectangle "Rectangle_5" at 195,48 size 29x9
      Visibility <- "DB_HMI_Start_System"
      Appearance <- "DB_HMI_Start_System"
   Button "Button_3" at 250,84 size 63x27; TextOff 'Set T=0C / Stellen T=0C'
      on Press: SetTag("DB_HMI_Set_T0", 1)
      on Release: SetTag("DB_HMI_Set_T0", 0)
   Button "Button_4" at 250,52 size 63x27; TextOff 'Set T=50C / Stellen Sie T=50C'
      on Release: SetTag("DB_HMI_Set_T50", 0)
      on Press: SetTag("DB_HMI_Set_T50", 1)
   Button "Button_5" at 176,154 size 135x49; TextOff 'Inspect Pistons Prüfen Kolben'
      on Press: ActivateScreen("Inspect Pistoane", 0)
*)

(* ===== HMI "HMI_RT_3" =====
system functions are stored by id; their names below are inferred from use
connection "HMI_Connection_4": ETHERNET, SIMATIC S7 300/400 MPI

HMI tags "Default tag table"
   "Emg_Stop_1" : Bool AT %I0.3, 100 ms
   "Automata" : UInt, internal
   "DB_SIM_BTN_RESET" : Bool = PLC DB_SIM.BTN_RESET AT %DB40.DBX0.4, 100 ms
   "Emg_Stop" : Bool = PLC Emg_Stop AT %I0.2, 100 ms
   "Final_Cursa_P1" : Bool = PLC Final_Cursa_Piston_1 AT %M2.5, 100 ms
   "Greutate" : Int AT %DB7.DBW2, 100 ms
   "LOAD" : Bool = PLC Banda_1_DB.Btn_LOAD AT %DB8.DBX0.4, 100 ms
   "Loc_Ocupat_A" : Int AT %DB1.DBW0, 100 ms
   "Locuri_A" : Int = PLC DB_HMI.Locuri_A AT %DB19.DBW0, 100 ms
   "Locuri_B" : Int = PLC DB_HMI.Locuri_B AT %DB19.DBW2, 100 ms
   "Locuri_C" : Int = PLC DB_HMI.Locuri_C AT %DB19.DBW4, 100 ms
   "Man/Auto" : Bool = PLC "Man/Auto" AT %I0.3, 100 ms
   "ON/OFF" : Bool = PLC "ON/OFF" AT %M2.1, 100 ms
   "Poz_Cutie" : Int = PLC Poz_Cutie AT %MW0, Cycle_1
   "Poz_Piston_1" : Int = PLC DB_general.Poz_Piston_1 AT %DB2.DBW2, Cycle_1
   "Start" : Bool = PLC Start AT %I0.0, 100 ms
   "StatieDistributie" : UInt, internal
   "StatieHidraulica" : UInt, internal
   "StatieIncarcare" : UInt, internal
   "Stop" : Bool = PLC Stop AT %I0.1, 100 ms
   "Tag_ScreenNumber" : UInt, internal
   "Viz_Cutie_Cursa_Scurta" : Bool = PLC Viz_Cutie_Cursa_Scurta AT %M2.2, 100 ms
   "RdyToLog" : Bool = PLC DB_InsertCutieTrigger.Readytolog AT %DB5.DBX8.0, 100 ms
      on ChangeValue: "VBFunction_4"()
   "Greutate_Pachet" : Int = PLC DB_InsertCutieTrigger.Greutate_Pachet AT %DB5.DBW12, 100 ms
   "Destinatie_Pachet" : Int = PLC DB_InsertCutieTrigger.Destinatie_Pachet AT %DB5.DBW10, 100 ms
   "Tip_Cutie_Pachet" : Int = PLC DB_InsertCutieTrigger.Tip_Cutie_Pachet AT %DB5.DBW14, 100 ms
   "Destinatie_1" : Int, internal
   "Tip_1" : Int, internal
   "Greutate_1" : Int, internal
   "Id_1" : Int, internal
   "url" : WString[254], internal
   "Data" : DateTime, internal
   "QR_TEST" : Bool, internal
   "ID_TEST" : Int, internal
   "Greutate_TEST" : Int, internal
   "Destinatie_TEST" : WString[254], internal
   "Tip_TEST" : WString[254], internal
   "Array_Id" : Array [0..10] of Int, internal
   "Array_Data" : Array [0..10] of DateTime, internal
   "DB_Tranzitii_Viz_Cutie_1" : Bool = PLC DB_Tranzitii.VizCutieStart AT %DB47.DBX0.0, 100 ms
   "DB_Tranzitii_Tip_Cutie_Man/Auto" : Int = PLC DB_Tranzitii.Tip_Cutie_Man/Auto_Start AT %DB47.DBW2, 100 ms
   "DB_Tranzitii_VizCutieEnd" : Bool = PLC DB_Tranzitii.VizCutieEnd AT %DB47.DBX4.0, 100 ms
   "DB_Tranzitii_TipCutieMan/Auto_End" : Int = PLC DB_Tranzitii.TipCutieMan/Auto_End AT %DB47.DBW6, 100 ms
   "DB_Vizibilitati_Platforme/Colete_Platforma_A" : Bool = PLC "DB_Vizibilitati_Platforme/Colete".Platforma_A AT %DB1.DBX0.0, 100 ms
   "DB_Vizibilitati_Platforme/Colete_Colet_A" : Bool = PLC "DB_Vizibilitati_Platforme/Colete".Colet_A AT %DB1.DBX0.3, 100 ms
   "DB_RemoteAcces_EmgStopBtn" : Bool = PLC DB_general.Stare_Poz_Incarcare AT %DB6.DBX0.0, 100 ms
   "DB_RemoteAcces_Stop" : Bool = PLC DB_general.Poz_Piston_1 AT %DB6.DBX0.1, 100 ms
   "DB_RemoteAcces_Start" : Bool = PLC DB_HMI.A_Pressed AT %DB6.DBX0.2, 100 ms
   "DB_RemoteAcces_Manual/Auto" : Bool = PLC DB_HMI.B_Pressed AT %DB6.DBX0.3, 100 ms
   "DB_RemoteAcces_On/Off" : Bool = PLC DB_HMI.C_Pressed AT %DB6.DBX0.4, 100 ms
   "DB_RemoteAcces_Remote" : Bool = PLC DB_HMI.Cutie_Manuala AT %DB6.DBX0.5, 100 ms
   "Data_Control_En_Load_Enable" : Bool = PLC DB_HMI.Cutie_Automata AT %DB14.DBX0.0, 1 s
   "DB_Vizibilitati_Platforme/Colete_Colet_B" : Bool = PLC DB_HMI.Viz_Cutie_Scurta AT %DB1.DBX0.4, 100 ms
   "DB_Vizibilitati_Platforme/Colete_Platforma_B" : Bool = PLC DB_general.Senzor_1_Incarcare AT %DB1.DBX0.1, 100 ms
   "DB_Vizibilitati_Platforme/Colete_Platforma_C" : Bool = PLC DB_general.Senzor_2_Incarcare AT %DB1.DBX0.2, 100 ms
   "DB_Vizibilitati_Platforme/Colete_Colet_C" : Bool = PLC DB_HMI.Tip_Cutie_Lung AT %DB1.DBX0.5, 100 ms
   "DB_general_GreutateManual" : Real = PLC DB_HMI.LOAD AT %DB2.DBD44, 1 s
   "DB_general_GreutateAutomata" : Real = PLC DB_HMI.Transport AT %DB2.DBD48, 1 s
   "DB_HMI_Detalii_Cutii" : Int = PLC DB_HMI.Viz_Cutie_Lunga AT %DB19.DBW70, 100 ms
   "DB_HMI_Modificare_Param" : Int = PLC DB_HMI.Packets_Param AT %DB19.DBW72, 1 s
   "DB_HMI_MaxLoad_A" : Int = PLC DB_HMI.MaxLoad_A AT %DB19.DBW74, 1 s
   "DB_HMI_MaxLoad_B" : Int = PLC DB_general.Senzor_1_Descarcare AT %DB19.DBW76, 1 s
   "DB_HMI_MaxLoad_C" : Int = PLC DB_general.Valoare AT %DB19.DBW78, 1 s
   "DB_HMI_Cantitate_A" : Int = PLC DB_HMI.Cantitate_A AT %DB19.DBW80, 1 s
   "DB_HMI_Cantitate_B" : Int = PLC DB_general.Piston_1_Cursa_Completa AT %DB19.DBW82, 1 s
   "DB_HMI_Cantitat_C" : Int = PLC DB_HMI.Viz_Cutie_Banda_1 AT %DB19.DBW84, 1 s
   "DB_HMI_Pachete_Schimb1" : Int = PLC DB_HMI.Ack_Load AT %DB19.DBW88, 1 s
   "DB_HMI_Pachete_Schimb2" : Int = PLC DB_HMI.Piston_1_Status AT %DB19.DBW90, 1 s
   "DB_HMI_Pachete_Schimb3" : Int = PLC DB_HMI.Piston_2_Status AT %DB19.DBW92, 1 s
   "DB_HMI_Total_Packets" : Int = PLC DB_general.Piston_2_Cursa_Completa AT %DB19.DBW86, 1 s
   "DB_HMI_Sistem_Racire" : Bool = PLC DB_HMI.Load_RDY AT %DB19.DBX94.0, 1 s
   "DB_HMI_Temp_Min" : Int = PLC DB_general.Poz_Cutie_Bile AT %DB19.DBW98, 1 s
   "DB_HMI_Temp_Max" : Int = PLC DB_HMI.Viz_Cutie_A AT %DB19.DBW96, 1 s
   "DB_HMI_Temp_Optim" : Int = PLC DB_HMI.Viz_Cutie_B AT %DB19.DBW100, 1 s
   "DB_general_Procent_Toleranta" : Real = PLC DB_HMI.Viz_Cutie_C AT %DB2.DBD52, 1 s
   "DB_HMI_Detalii_Truck_A" : Bool = PLC DB_HMI.LOAD_A AT %DB19.DBX120.0, 100 ms
   "DB_HMI_Detalii_Truck_B" : Bool = PLC DB_general.Piston_Incarcare_A AT %DB19.DBX120.1, 100 ms
   "DB_HMI_Detalii_Truck_C" : Bool = PLC DB_HMI.LOAD_B AT %DB19.DBX120.2, 100 ms
   "DB_HMI_Cantitate_Loaded_B" : Int = PLC DB_HMI.LOAD_C AT %DB19.DBW116, 1 s
   "DB_HMI_Total_Weight_B" : Real = PLC DB_general.Piston_Incarcare_B AT %DB19.DBD106, 1 s
   "DB_HMI_Cantitate_Loaded_C" : Int = PLC DB_general.Piston_Incarcare_C AT %DB19.DBW118, 1 s
   "DB_HMI_Total_Weight_C" : Real = PLC DB_HMI.Status_Piston_A AT %DB19.DBD110, 1 s
   "DB_HMI_Cantitate_Loaded_A" : Int = PLC DB_HMI.Status_Piston_B AT %DB19.DBW114, 1 s
   "DB_HMI_Total_Weight_A" : Real = PLC DB_HMI.Status_Piston_C AT %DB19.DBD102, 1 s
   "Template_Satie_Distribuire" : Bool = PLC DB_HMI.Status_Banda_Bile AT %DB16.DBX0.0, 1 s
   "Template_Statie_Incarcare" : Bool = PLC DB_HMI.Sageata_Deplasare_Banda_Bile AT %DB16.DBX0.1, 1 s
   "Template_Packets_Log" : Bool = PLC DB_HMI.Temp_Ulei AT %DB16.DBX0.2, 1 s
   "Template_Hidraulic_Station" : Bool = PLC DB_HMI.Volum_Ulei AT %DB16.DBX0.3, 1 s
   "Template_Errors" : Bool = PLC DB_HMI.Add_Ulei AT %DB16.DBX0.4, 1 s
   "Template_Home" : Bool = PLC DB_HMI.Sub_Ulei AT %DB16.DBX0.5, 1 s
   "DB_general_GreutateMaxManual" : Real = PLC DB_HMI.Tip_Cutie_Scurt AT %DB2.DBD72, 1 s
   "DB_general_GreutateMinAutomat" : Real = PLC DB_HMI.Start_System AT %DB2.DBD76, 1 s
   "DB_Tip_Cutie_GreutateCutie" : Real = PLC DB_HMI.Racire_Ulei AT %DB37.DBD0, 1 s
   "DB_Tip_Cutie_IntersectieInterval" : Int = PLC DB_HMI.Set_T0 AT %DB37.DBW4, 1 s
   "DB_Tip_Cutie_TipCutie" : Bool = PLC DB_HMI.Set_T50 AT %DB37.DBX6.0, 100 ms
   "DB_Tip_Cutie_VizTipCutie" : Bool = PLC DB_HMI.START_SIM AT %DB37.DBX6.1, 100 ms
   "DB_general_GreutateMinManual" : Real = PLC DB_HMI.BTN_LOAD AT %DB2.DBD68, 1 s
   "DB_general_GreutateMaxAutomat" : Real = PLC DB_Alarme.Emg_Stop AT %DB2.DBD80, 1 s
   "DB_Tip_Cutie_RebutLbl" : Bool = PLC DB_HMI.Status_Incalzire/Racire_Ulei AT %DB37.DBX6.2, 100 ms
   "DB_Tip_Cutie_Scrap" : Int = PLC DB_HMI.Viz_Cutie_Man/Auto AT %DB37.DBW8, 100 ms
   "DB_Inspect_Pistoane_PompaPrincipala" : Int = PLC DB_HMI.Ventilator_Rece AT %DB34.DBW20, 1 s
   "DB_Inspect_Pistoane_Pompa1" : Int = PLC DB_HMI.Ventilator_Cald AT %DB34.DBW22, 1 s
   "DB_Inspect_Pistoane_Pompa2" : Int = PLC DB_Inspect_Pistoane.Piston_1 AT %DB34.DBW24, 1 s
   "DB_Inspect_Pistoane_PompaA" : Int = PLC DB_Inspect_Pistoane.Piston_2 AT %DB34.DBW26, 1 s